(* Logix 5000 project; controller PLC_MCC1201_220AP1 vendor 1 type 14 code 164 rev 35.11; software revision 35.00; part 10 of 25 *)
(* tags used below, declared in another part *)
   TMP_rDummy : REAL;
   TMP_rTarget : REAL;
   TMP_xDummy : BOOL;
   B3 : DINT[102];
   GP_OB_InitializeMain : GP_OB_Initialize;
   HMI_Alarm_Reset : BOOL;   // HMI_Alarm_Reset
   HMI_MAN_CMD_WR : UDT_MAN_CMD_WR;
   LEHR_SPEED : ALIAS FOR N60[1];
   M225 : MAC_EMERGENCYXCUT;
   M225_HMW : MAC_EMERGENCYXCUT_HMW;
   M225_M1_DR : AXIS_CIP_DRIVE;
   M225_OUT_MOTION : MAC_EMERGENCYXCUT_OUT_MOTION;
   M2xx_CONVEYOR : MAC_CONVEYOR[20];
   M2xx_CONVEYOR_IN_MOTION : MAC_CONVEYOR_IN_MOTION[20];
   M2xx_CONVEYOR_OUT_MOTION : MAC_CONVEYOR_OUT_MOTION[20];
   M301_M1_DR : AXIS_CIP_DRIVE;
   M301_M2_DR : AXIS_CIP_DRIVE;
   TMP_dDirection : DINT;
   TMP_rAcc : REAL;
   TMP_rDec : REAL;
   TMP_rSpeed : REAL;
   TMP_xAlwaysOFF : BOOL;
   TMP_xRun : BOOL;
   Z200_UPS : ZONE_UPS;
(* CommandLogic, continued *)

ROUTINE M225_EmergencyCut_Outputs   (* ladder *)
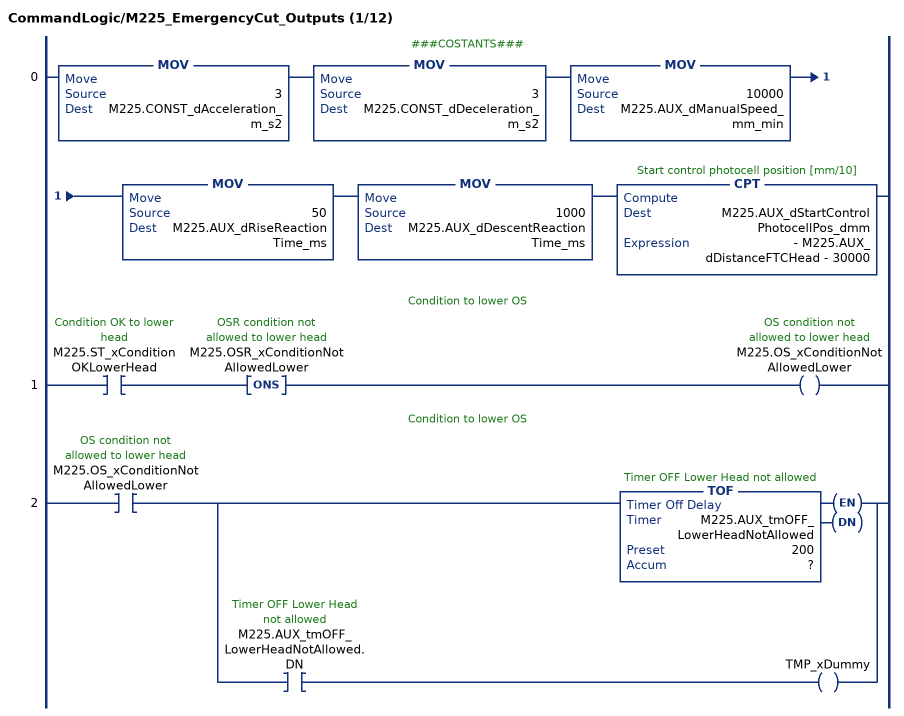
   // ###COSTANTS###
   0: MOV(3,M225.CONST_dAcceleration_m_s2)MOV(3,M225.CONST_dDeceleration_m_s2)MOV(10000,M225.AUX_dManualSpeed_mm_min)MOV(50,M225.AUX_dRiseReactionTime_ms)MOV(1000,M225.AUX_dDescentReactionTime_ms)CPT(M225.AUX_dStartControlPhotocellPos_dmm,- M225.AUX_dDistanceFTCHead - 30000);
   // Condition to lower OS
   1: XIC(M225.ST_xConditionOKLowerHead)ONS(M225.OSR_xConditionNotAllowedLower)OTE(M225.OS_xConditionNotAllowedLower);
   // Condition to lower OS
   2: XIC(M225.OS_xConditionNotAllowedLower)[TOF(M225.AUX_tmOFF_LowerHeadNotAllowed,?,?) ,XIC(M225.AUX_tmOFF_LowerHeadNotAllowed.DN) OTE(TMP_xDummy) ];
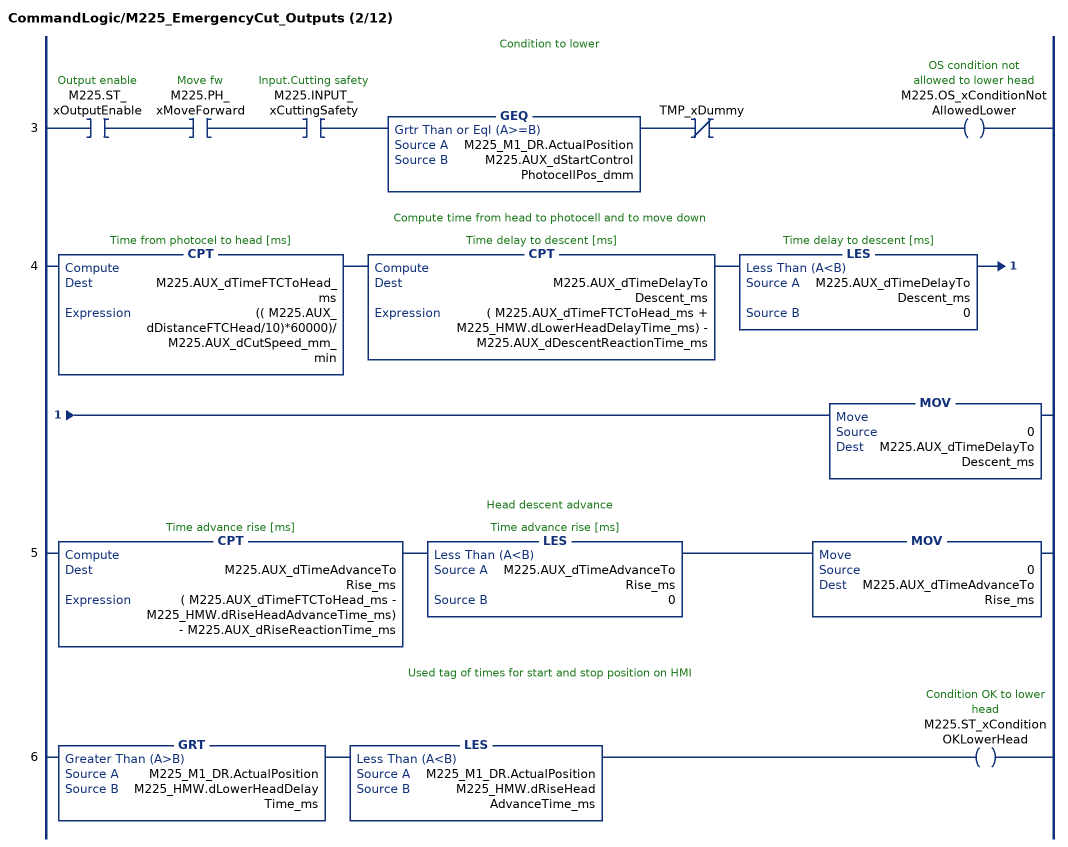
   // Condition to lower
   3: XIC(M225.ST_xOutputEnable)XIC(M225.PH_xMoveForward)XIC(M225.INPUT_xCuttingSafety)GEQ(M225_M1_DR.ActualPosition,M225.AUX_dStartControlPhotocellPos_dmm)XIO(TMP_xDummy)OTE(M225.OS_xConditionNotAllowedLower);
   // Compute time from head to photocell and to move down
   4: CPT(M225.AUX_dTimeFTCToHead_ms,(( M225.AUX_dDistanceFTCHead/10)*60000)/ M225.AUX_dCutSpeed_mm_min)CPT(M225.AUX_dTimeDelayToDescent_ms,( M225.AUX_dTimeFTCToHead_ms + M225_HMW.dLowerHeadDelayTime_ms) - M225.AUX_dDescentReactionTime_ms)LES(M225.AUX_dTimeDelayToDescent_ms,0)MOV(0,M225.AUX_dTimeDelayToDescent_ms);
   // Head descent advance
   5: CPT(M225.AUX_dTimeAdvanceToRise_ms,( M225.AUX_dTimeFTCToHead_ms - M225_HMW.dRiseHeadAdvanceTime_ms) - M225.AUX_dRiseReactionTime_ms)LES(M225.AUX_dTimeAdvanceToRise_ms,0)MOV(0,M225.AUX_dTimeAdvanceToRise_ms);
   // Used tag of times for start and stop position on HMI
   6: GRT(M225_M1_DR.ActualPosition,M225_HMW.dLowerHeadDelayTime_ms)LES(M225_M1_DR.ActualPosition,M225_HMW.dRiseHeadAdvanceTime_ms)OTE(M225.ST_xConditionOKLowerHead);
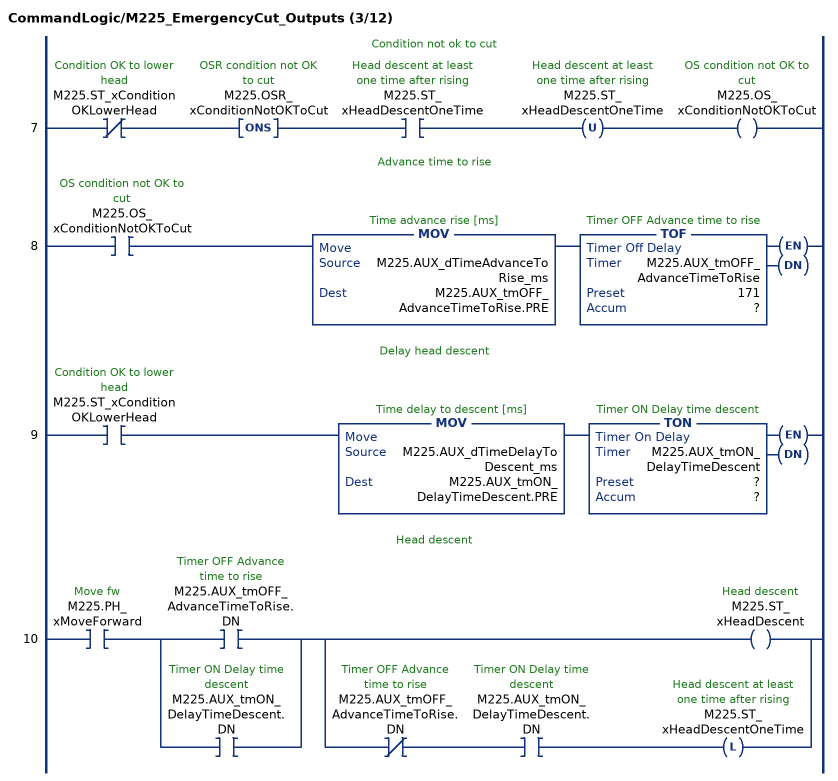
   // Condition not ok to cut
   7: XIO(M225.ST_xConditionOKLowerHead)ONS(M225.OSR_xConditionNotOKToCut)XIC(M225.ST_xHeadDescentOneTime)OTU(M225.ST_xHeadDescentOneTime)OTE(M225.OS_xConditionNotOKToCut);
   // Advance time to rise
   8: XIC(M225.OS_xConditionNotOKToCut)MOV(M225.AUX_dTimeAdvanceToRise_ms,M225.AUX_tmOFF_AdvanceTimeToRise.PRE)TOF(M225.AUX_tmOFF_AdvanceTimeToRise,?,?);
   // Delay head descent
   9: XIC(M225.ST_xConditionOKLowerHead)MOV(M225.AUX_dTimeDelayToDescent_ms,M225.AUX_tmON_DelayTimeDescent.PRE)TON(M225.AUX_tmON_DelayTimeDescent,?,?);
   // Head descent
   10: XIC(M225.PH_xMoveForward)[XIC(M225.AUX_tmOFF_AdvanceTimeToRise.DN) ,XIC(M225.AUX_tmON_DelayTimeDescent.DN) ][OTE(M225.ST_xHeadDescent) ,XIO(M225.AUX_tmOFF_AdvanceTimeToRise.DN) XIC(M225.AUX_tmON_DelayTimeDescent.DN) OTL(M225.ST_xHeadDescentOneTime) ];
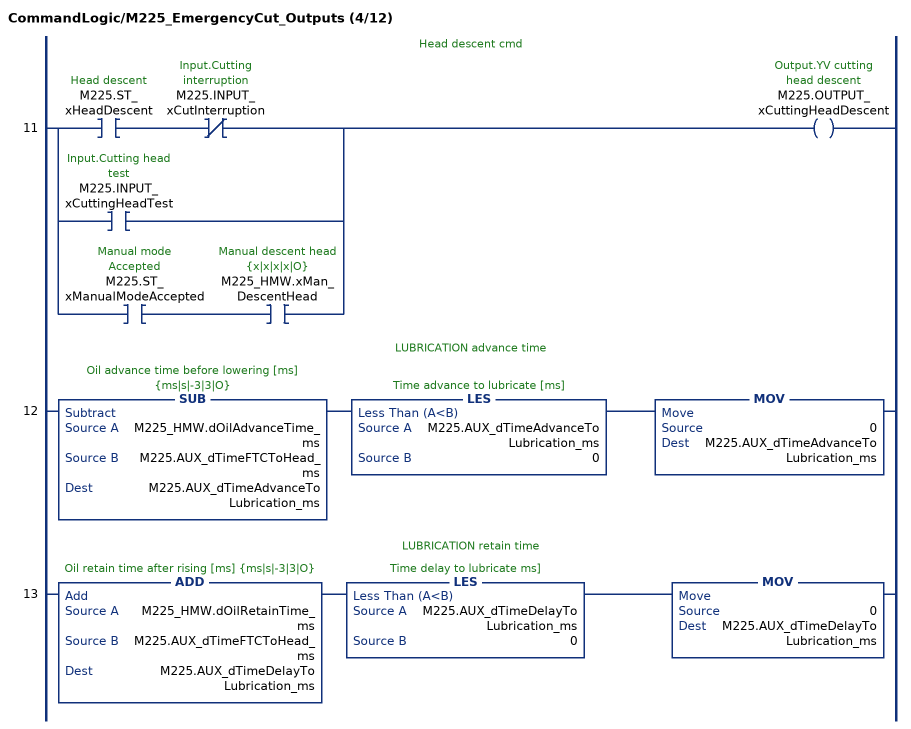
   // Head descent cmd
   11: [XIC(M225.ST_xHeadDescent) XIO(M225.INPUT_xCutInterruption) ,XIC(M225.INPUT_xCuttingHeadTest) ,XIC(M225.ST_xManualModeAccepted) XIC(M225_HMW.xMan_DescentHead) ]OTE(M225.OUTPUT_xCuttingHeadDescent);
   // LUBRICATION advance time
   12: SUB(M225_HMW.dOilAdvanceTime_ms,M225.AUX_dTimeFTCToHead_ms,M225.AUX_dTimeAdvanceToLubrication_ms)LES(M225.AUX_dTimeAdvanceToLubrication_ms,0)MOV(0,M225.AUX_dTimeAdvanceToLubrication_ms);
   // LUBRICATION retain time
   13: ADD(M225_HMW.dOilRetainTime_ms,M225.AUX_dTimeFTCToHead_ms,M225.AUX_dTimeDelayToLubrication_ms)LES(M225.AUX_dTimeDelayToLubrication_ms,0)MOV(0,M225.AUX_dTimeDelayToLubrication_ms);
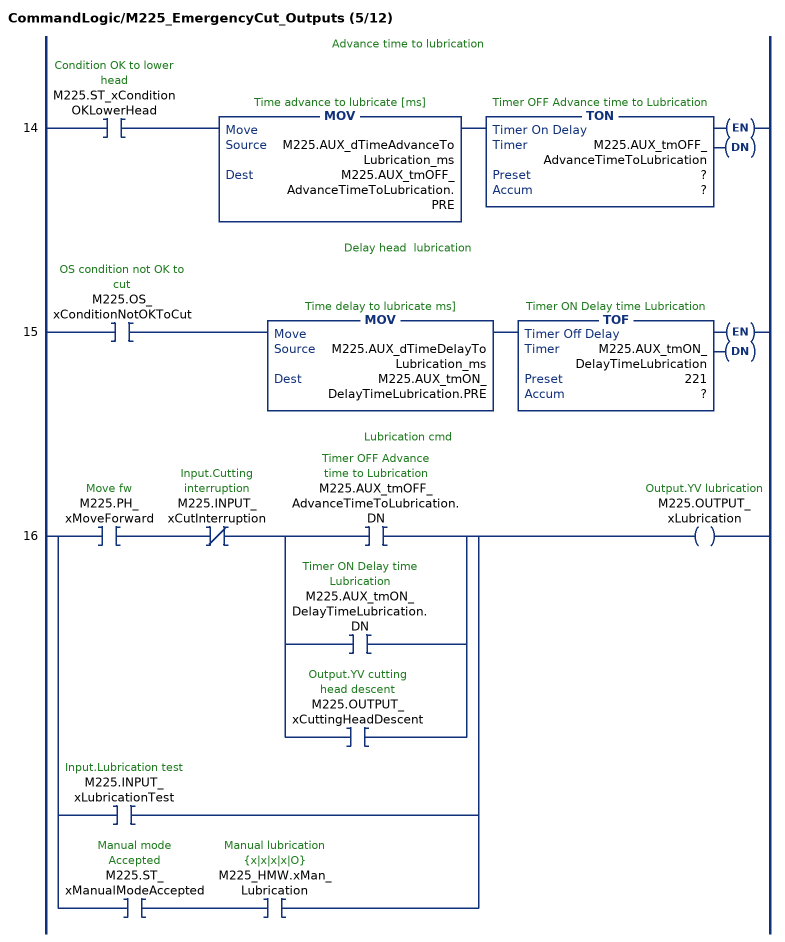
   // Advance time to lubrication
   14: XIC(M225.ST_xConditionOKLowerHead)MOV(M225.AUX_dTimeAdvanceToLubrication_ms,M225.AUX_tmOFF_AdvanceTimeToLubrication.PRE)TON(M225.AUX_tmOFF_AdvanceTimeToLubrication,?,?);
   // Delay head  lubrication
   15: XIC(M225.OS_xConditionNotOKToCut)MOV(M225.AUX_dTimeDelayToLubrication_ms,M225.AUX_tmON_DelayTimeLubrication.PRE)TOF(M225.AUX_tmON_DelayTimeLubrication,?,?);
   // Lubrication cmd
   16: [XIC(M225.PH_xMoveForward) XIO(M225.INPUT_xCutInterruption) [XIC(M225.AUX_tmOFF_AdvanceTimeToLubrication.DN) ,XIC(M225.AUX_tmON_DelayTimeLubrication.DN) ,XIC(M225.OUTPUT_xCuttingHeadDescent) ] ,XIC(M225.INPUT_xLubricationTest) ,XIC(M225.ST_xManualModeAccepted) XIC(M225_HMW.xMan_Lubrication) ]OTE(M225.OUTPUT_xLubrication);
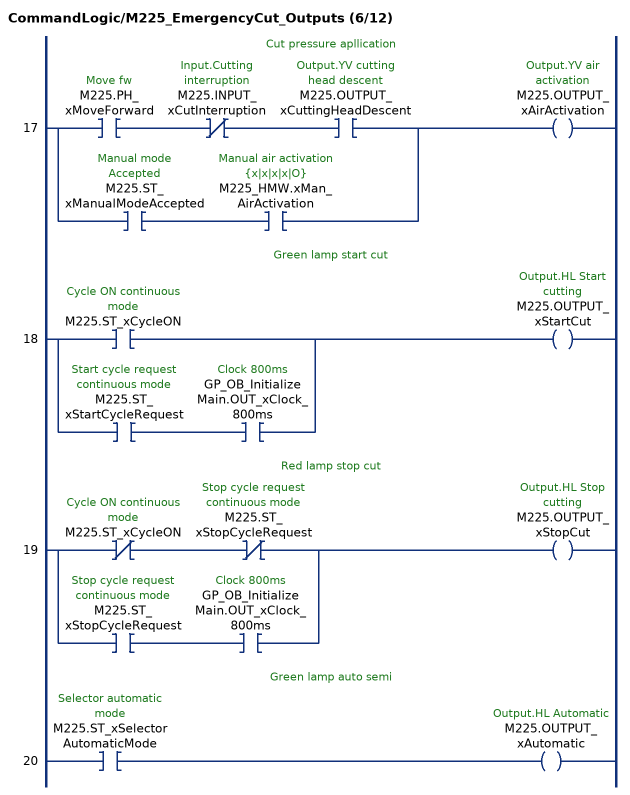
   // Cut pressure apllication
   17: [XIC(M225.PH_xMoveForward) XIO(M225.INPUT_xCutInterruption) XIC(M225.OUTPUT_xCuttingHeadDescent) ,XIC(M225.ST_xManualModeAccepted) XIC(M225_HMW.xMan_AirActivation) ]OTE(M225.OUTPUT_xAirActivation);
   // Green lamp start cut
   18: [XIC(M225.ST_xCycleON) ,XIC(M225.ST_xStartCycleRequest) XIC(GP_OB_InitializeMain.OUT_xClock_800ms) ]OTE(M225.OUTPUT_xStartCut);
   // Red lamp stop cut
   19: [XIO(M225.ST_xCycleON) XIO(M225.ST_xStopCycleRequest) ,XIC(M225.ST_xStopCycleRequest) XIC(GP_OB_InitializeMain.OUT_xClock_800ms) ]OTE(M225.OUTPUT_xStopCut);
   // Green lamp auto semi
   20: XIC(M225.ST_xSelectorAutomaticMode)OTE(M225.OUTPUT_xAutomatic);
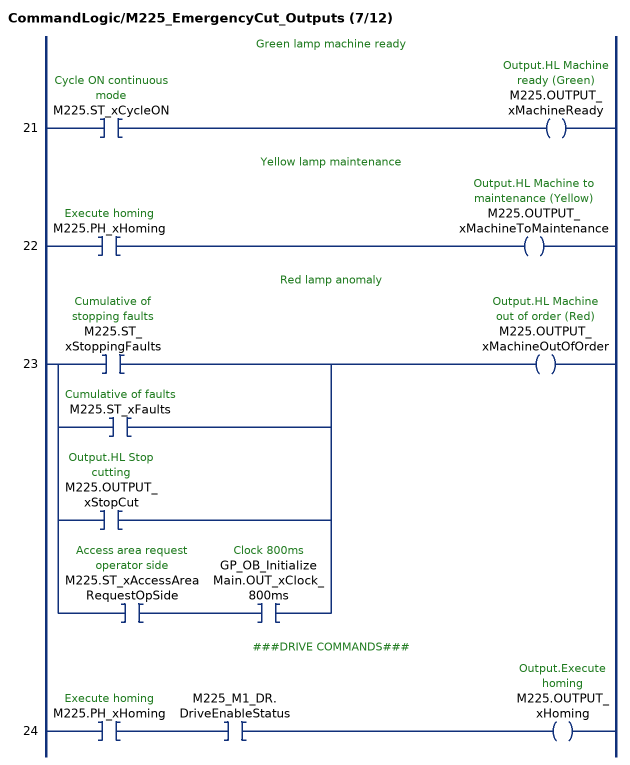
   // Green lamp machine ready
   21: XIC(M225.ST_xCycleON)OTE(M225.OUTPUT_xMachineReady);
   // Yellow lamp maintenance
   22: XIC(M225.PH_xHoming)OTE(M225.OUTPUT_xMachineToMaintenance);
   // Red lamp anomaly
   23: [XIC(M225.ST_xStoppingFaults) ,XIC(M225.ST_xFaults) ,XIC(M225.OUTPUT_xStopCut) ,XIC(M225.ST_xAccessAreaRequestOpSide) XIC(GP_OB_InitializeMain.OUT_xClock_800ms) ]OTE(M225.OUTPUT_xMachineOutOfOrder);
   // ###DRIVE COMMANDS###
   24: XIC(M225.PH_xHoming)XIC(M225_M1_DR.DriveEnableStatus)OTE(M225.OUTPUT_xHoming);
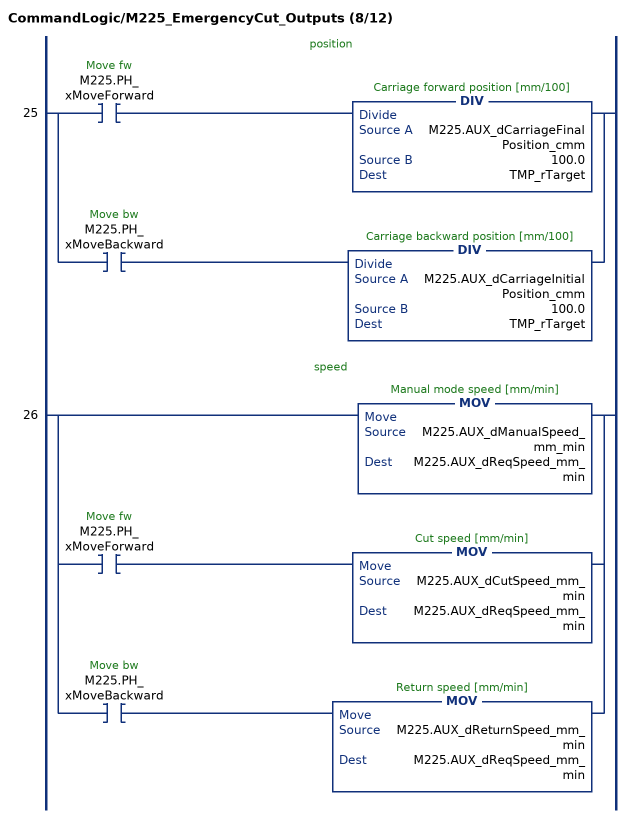
   // position
   25: [XIC(M225.PH_xMoveForward) DIV(M225.AUX_dCarriageFinalPosition_cmm,100.0,TMP_rTarget) ,XIC(M225.PH_xMoveBackward) DIV(M225.AUX_dCarriageInitialPosition_cmm,100.0,TMP_rTarget) ];
   // speed
   26: [MOV(M225.AUX_dManualSpeed_mm_min,M225.AUX_dReqSpeed_mm_min) ,XIC(M225.PH_xMoveForward) MOV(M225.AUX_dCutSpeed_mm_min,M225.AUX_dReqSpeed_mm_min) ,XIC(M225.PH_xMoveBackward) MOV(M225.AUX_dReturnSpeed_mm_min,M225.AUX_dReqSpeed_mm_min) ];
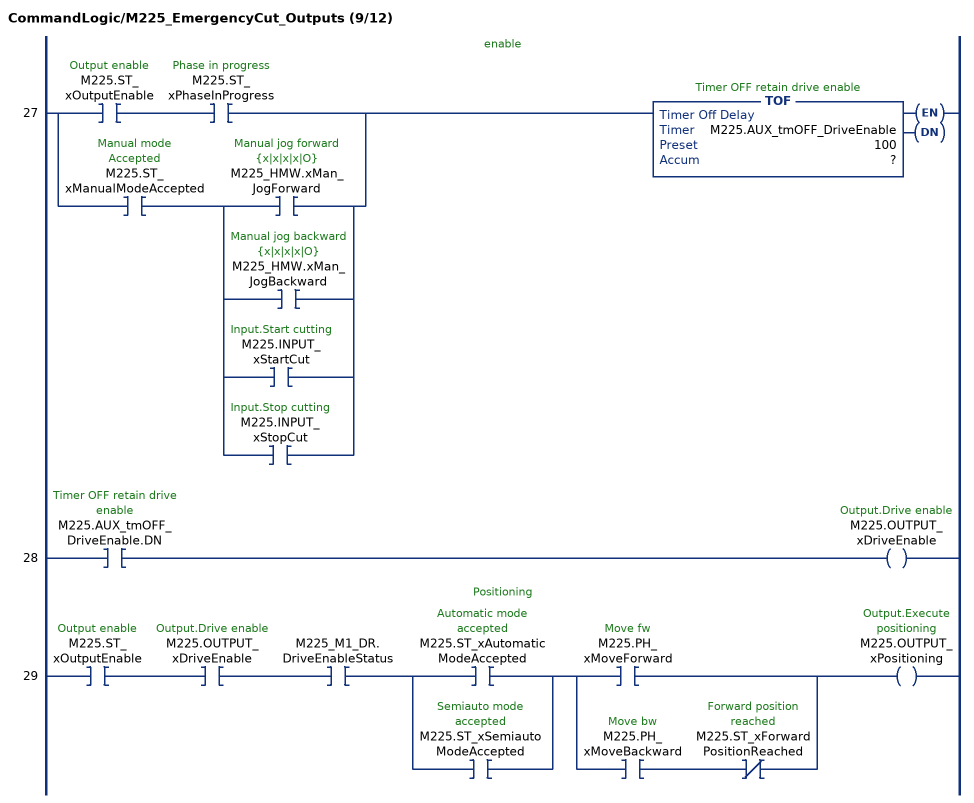
   // enable
   27: [XIC(M225.ST_xOutputEnable) XIC(M225.ST_xPhaseInProgress) ,XIC(M225.ST_xManualModeAccepted) [XIC(M225_HMW.xMan_JogForward) ,XIC(M225_HMW.xMan_JogBackward) ,XIC(M225.INPUT_xStartCut) ,XIC(M225.INPUT_xStopCut) ] ]TOF(M225.AUX_tmOFF_DriveEnable,?,?);
   28: XIC(M225.AUX_tmOFF_DriveEnable.DN)OTE(M225.OUTPUT_xDriveEnable);
   // Positioning
   29: XIC(M225.ST_xOutputEnable)XIC(M225.OUTPUT_xDriveEnable)XIC(M225_M1_DR.DriveEnableStatus)[XIC(M225.ST_xAutomaticModeAccepted) ,XIC(M225.ST_xSemiautoModeAccepted) ][XIC(M225.PH_xMoveForward) ,XIC(M225.PH_xMoveBackward) XIO(M225.ST_xForwardPositionReached) ]OTE(M225.OUTPUT_xPositioning);
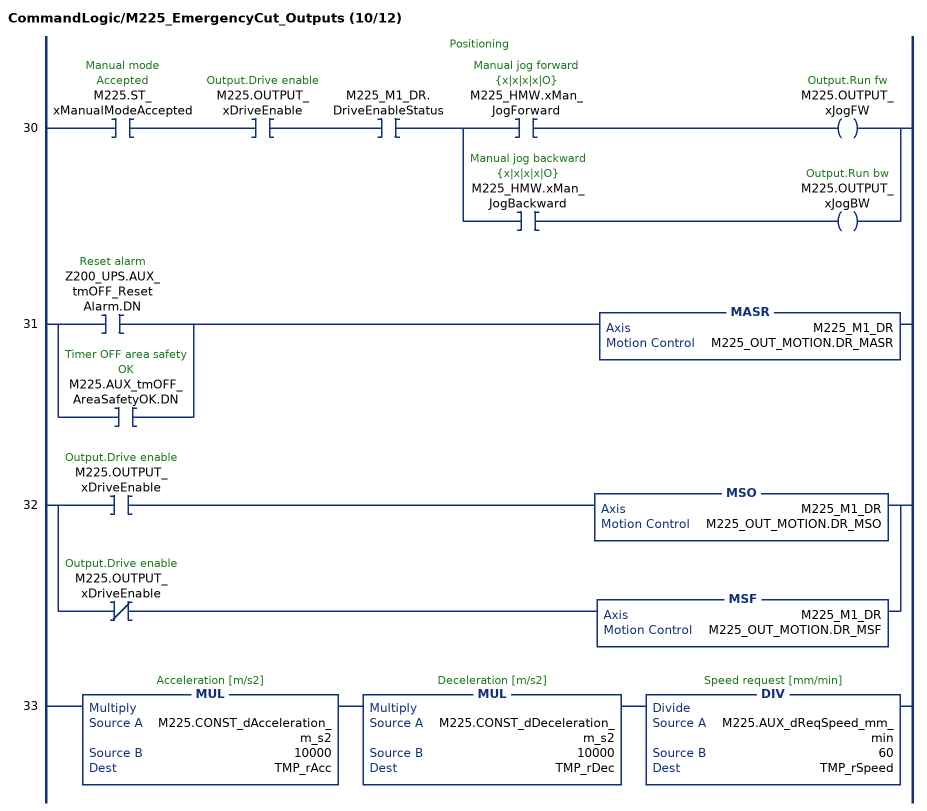
   // Positioning
   30: XIC(M225.ST_xManualModeAccepted)XIC(M225.OUTPUT_xDriveEnable)XIC(M225_M1_DR.DriveEnableStatus)[XIC(M225_HMW.xMan_JogForward) OTE(M225.OUTPUT_xJogFW) ,XIC(M225_HMW.xMan_JogBackward) OTE(M225.OUTPUT_xJogBW) ];
   31: [XIC(Z200_UPS.AUX_tmOFF_ResetAlarm.DN) ,XIC(M225.AUX_tmOFF_AreaSafetyOK.DN) ]MASR(M225_M1_DR,M225_OUT_MOTION.DR_MASR);
   32: [XIC(M225.OUTPUT_xDriveEnable) MSO(M225_M1_DR,M225_OUT_MOTION.DR_MSO) ,XIO(M225.OUTPUT_xDriveEnable) MSF(M225_M1_DR,M225_OUT_MOTION.DR_MSF) ];
   33: MUL(M225.CONST_dAcceleration_m_s2,10000,TMP_rAcc)MUL(M225.CONST_dDeceleration_m_s2,10000,TMP_rDec)DIV(M225.AUX_dReqSpeed_mm_min,60,TMP_rSpeed);
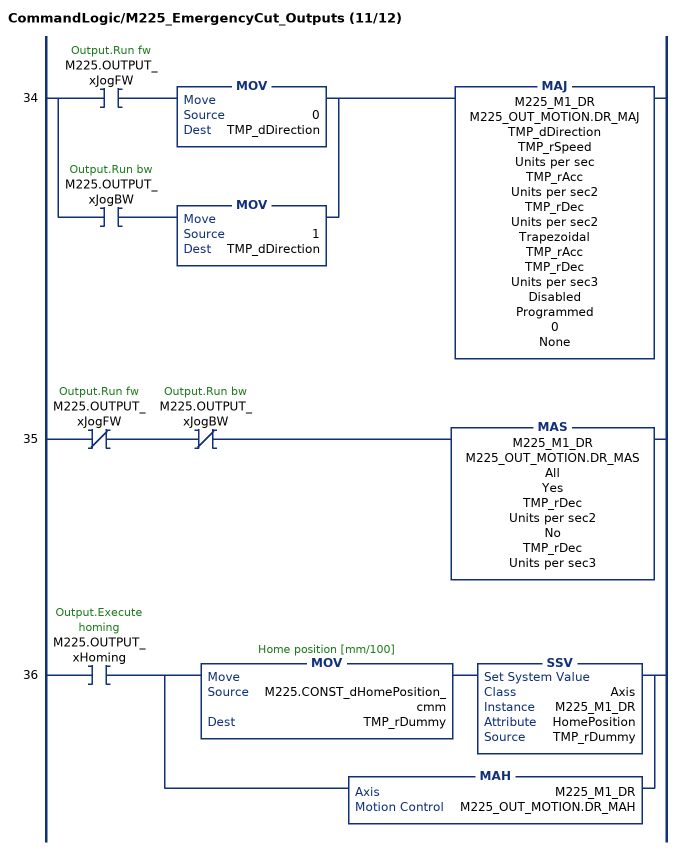
   34: [XIC(M225.OUTPUT_xJogFW) MOV(0,TMP_dDirection) ,XIC(M225.OUTPUT_xJogBW) MOV(1,TMP_dDirection) ]MAJ(M225_M1_DR,M225_OUT_MOTION.DR_MAJ,TMP_dDirection,TMP_rSpeed,Units per sec,TMP_rAcc,Units per sec2,TMP_rDec,Units per sec2,Trapezoidal,TMP_rAcc,TMP_rDec,Units per sec3,Disabled,Programmed,0,None);
   35: XIO(M225.OUTPUT_xJogFW)XIO(M225.OUTPUT_xJogBW)MAS(M225_M1_DR,M225_OUT_MOTION.DR_MAS,All,Yes,TMP_rDec,Units per sec2,No,TMP_rDec,Units per sec3);
   36: XIC(M225.OUTPUT_xHoming)[MOV(M225.CONST_dHomePosition_cmm,TMP_rDummy) SSV(Axis,M225_M1_DR,HomePosition,TMP_rDummy) ,MAH(M225_M1_DR,M225_OUT_MOTION.DR_MAH) ];
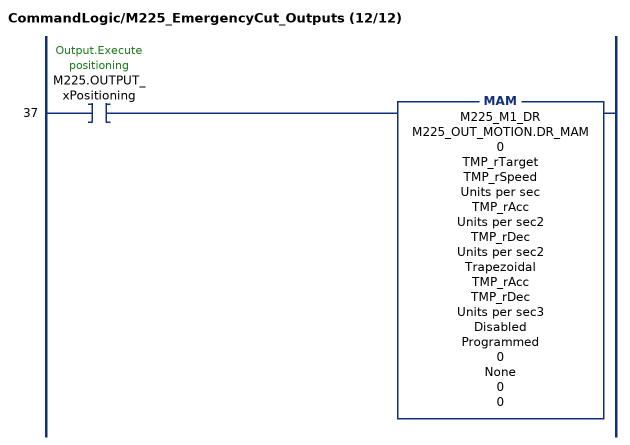
   37: XIC(M225.OUTPUT_xPositioning)MAM(M225_M1_DR,M225_OUT_MOTION.DR_MAM,0,TMP_rTarget,TMP_rSpeed,Units per sec,TMP_rAcc,Units per sec2,TMP_rDec,Units per sec2,Trapezoidal,TMP_rAcc,TMP_rDec,Units per sec3,Disabled,Programmed,0,None,0,0);
END_ROUTINE

ROUTINE M301M1_Conveyor_Motion_Output   (* ladder *)
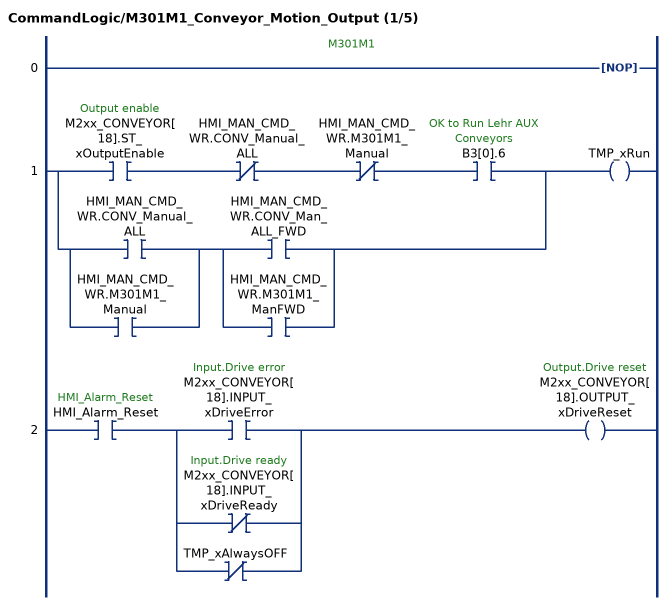
   // M301M1
   0: NOP();
   1: [XIC(M2xx_CONVEYOR[18].ST_xOutputEnable) XIO(HMI_MAN_CMD_WR.CONV_Manual_ALL) XIO(HMI_MAN_CMD_WR.M301M1_Manual) XIC(B3[0].6) ,[XIC(HMI_MAN_CMD_WR.CONV_Manual_ALL) ,XIC(HMI_MAN_CMD_WR.M301M1_Manual) ] [XIC(HMI_MAN_CMD_WR.CONV_Man_ALL_FWD) ,XIC(HMI_MAN_CMD_WR.M301M1_ManFWD) ] ]OTE(TMP_xRun);
   2: XIC(HMI_Alarm_Reset)[XIC(M2xx_CONVEYOR[18].INPUT_xDriveError) ,XIO(M2xx_CONVEYOR[18].INPUT_xDriveReady) ,XIO(TMP_xAlwaysOFF) ]OTE(M2xx_CONVEYOR[18].OUTPUT_xDriveReset);
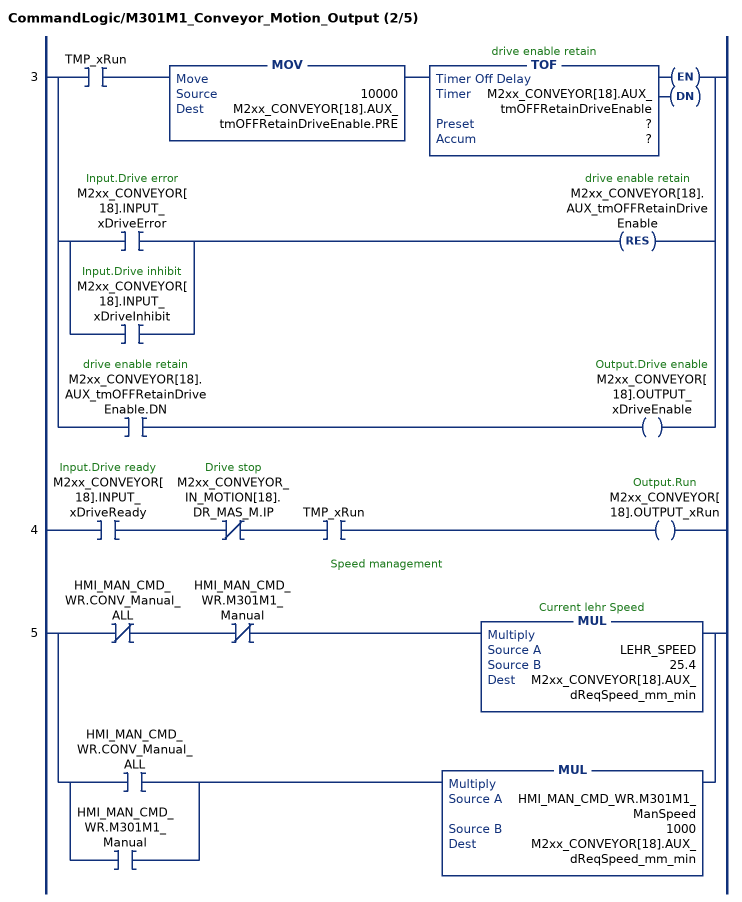
   3: [XIC(TMP_xRun) MOV(10000,M2xx_CONVEYOR[18].AUX_tmOFFRetainDriveEnable.PRE) TOF(M2xx_CONVEYOR[18].AUX_tmOFFRetainDriveEnable,?,?) ,[XIC(M2xx_CONVEYOR[18].INPUT_xDriveError) ,XIC(M2xx_CONVEYOR[18].INPUT_xDriveInhibit) ] RES(M2xx_CONVEYOR[18].AUX_tmOFFRetainDriveEnable) ,XIC(M2xx_CONVEYOR[18].AUX_tmOFFRetainDriveEnable.DN) OTE(M2xx_CONVEYOR[18].OUTPUT_xDriveEnable) ];
   4: XIC(M2xx_CONVEYOR[18].INPUT_xDriveReady)XIO(M2xx_CONVEYOR_IN_MOTION[18].DR_MAS_M.IP)XIC(TMP_xRun)OTE(M2xx_CONVEYOR[18].OUTPUT_xRun);
   // Speed management
   5: [XIO(HMI_MAN_CMD_WR.CONV_Manual_ALL) XIO(HMI_MAN_CMD_WR.M301M1_Manual) MUL(LEHR_SPEED,25.4,M2xx_CONVEYOR[18].AUX_dReqSpeed_mm_min) ,[XIC(HMI_MAN_CMD_WR.CONV_Manual_ALL) ,XIC(HMI_MAN_CMD_WR.M301M1_Manual) ] MUL(HMI_MAN_CMD_WR.M301M1_ManSpeed,1000,M2xx_CONVEYOR[18].AUX_dReqSpeed_mm_min) ];
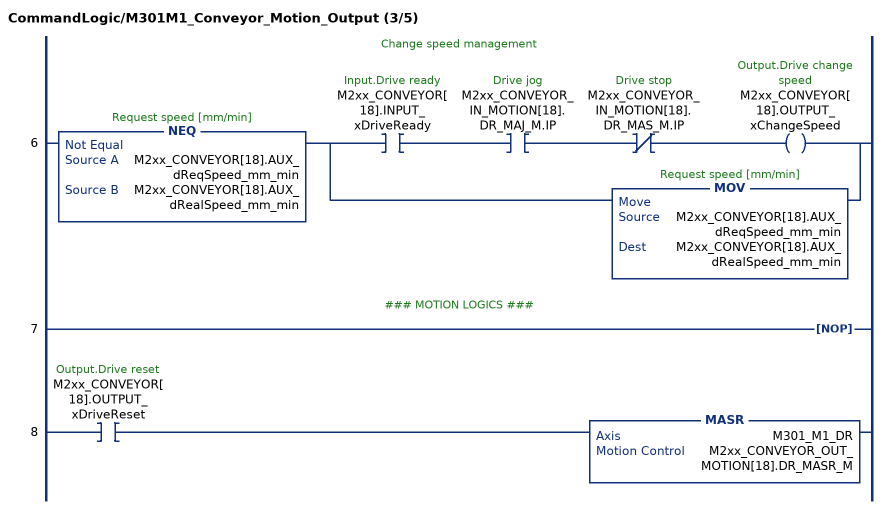
   // Change speed management
   6: NEQ(M2xx_CONVEYOR[18].AUX_dReqSpeed_mm_min,M2xx_CONVEYOR[18].AUX_dRealSpeed_mm_min)[XIC(M2xx_CONVEYOR[18].INPUT_xDriveReady) XIC(M2xx_CONVEYOR_IN_MOTION[18].DR_MAJ_M.IP) XIO(M2xx_CONVEYOR_IN_MOTION[18].DR_MAS_M.IP) OTE(M2xx_CONVEYOR[18].OUTPUT_xChangeSpeed) ,MOV(M2xx_CONVEYOR[18].AUX_dReqSpeed_mm_min,M2xx_CONVEYOR[18].AUX_dRealSpeed_mm_min) ];
   // ### MOTION LOGICS ###
   7: NOP();
   8: XIC(M2xx_CONVEYOR[18].OUTPUT_xDriveReset)MASR(M301_M1_DR,M2xx_CONVEYOR_OUT_MOTION[18].DR_MASR_M);
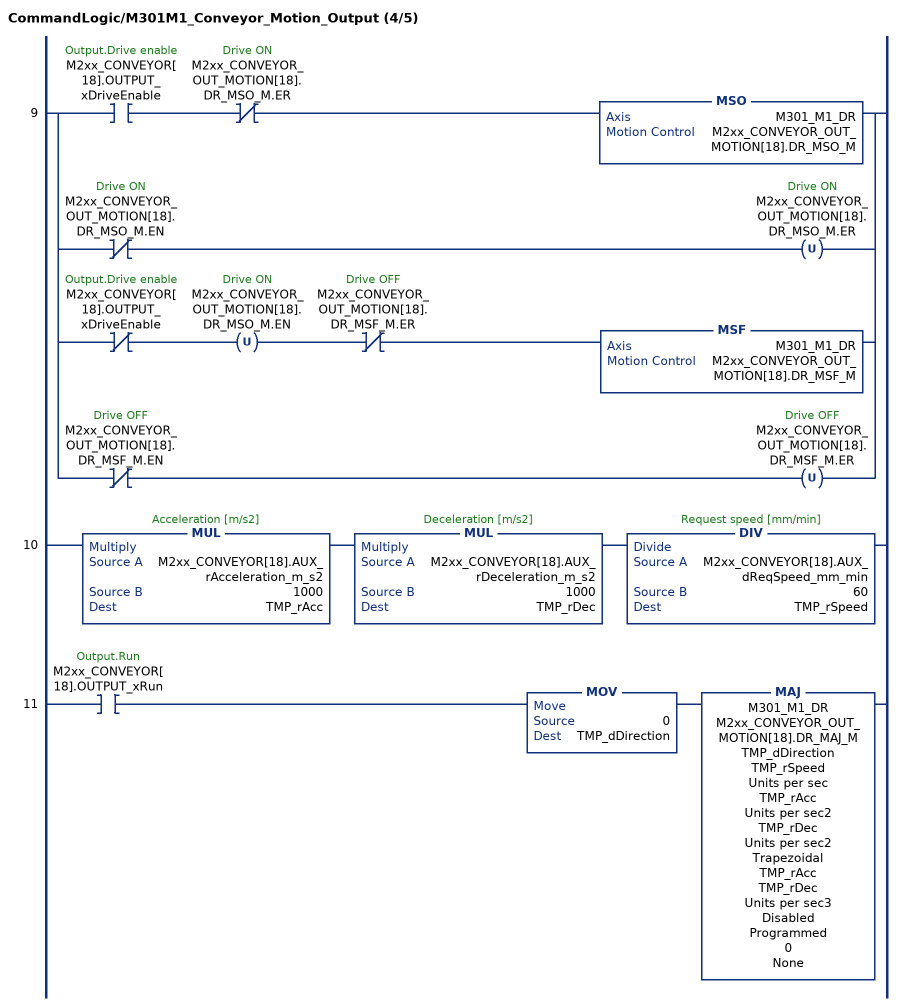
   9: [XIC(M2xx_CONVEYOR[18].OUTPUT_xDriveEnable) XIO(M2xx_CONVEYOR_OUT_MOTION[18].DR_MSO_M.ER) MSO(M301_M1_DR,M2xx_CONVEYOR_OUT_MOTION[18].DR_MSO_M) ,XIO(M2xx_CONVEYOR_OUT_MOTION[18].DR_MSO_M.EN) OTU(M2xx_CONVEYOR_OUT_MOTION[18].DR_MSO_M.ER) ,XIO(M2xx_CONVEYOR[18].OUTPUT_xDriveEnable) OTU(M2xx_CONVEYOR_OUT_MOTION[18].DR_MSO_M.EN) XIO(M2xx_CONVEYOR_OUT_MOTION[18].DR_MSF_M.ER) MSF(M301_M1_DR,M2xx_CONVEYOR_OUT_MOTION[18].DR_MSF_M) ,XIO(M2xx_CONVEYOR_OUT_MOTION[18].DR_MSF_M.EN) OTU(M2xx_CONVEYOR_OUT_MOTION[18].DR_MSF_M.ER) ];
   10: MUL(M2xx_CONVEYOR[18].AUX_rAcceleration_m_s2,1000,TMP_rAcc)MUL(M2xx_CONVEYOR[18].AUX_rDeceleration_m_s2,1000,TMP_rDec)DIV(M2xx_CONVEYOR[18].AUX_dReqSpeed_mm_min,60,TMP_rSpeed);
   11: XIC(M2xx_CONVEYOR[18].OUTPUT_xRun)MOV(0,TMP_dDirection)MAJ(M301_M1_DR,M2xx_CONVEYOR_OUT_MOTION[18].DR_MAJ_M,TMP_dDirection,TMP_rSpeed,Units per sec,TMP_rAcc,Units per sec2,TMP_rDec,Units per sec2,Trapezoidal,TMP_rAcc,TMP_rDec,Units per sec3,Disabled,Programmed,0,None);
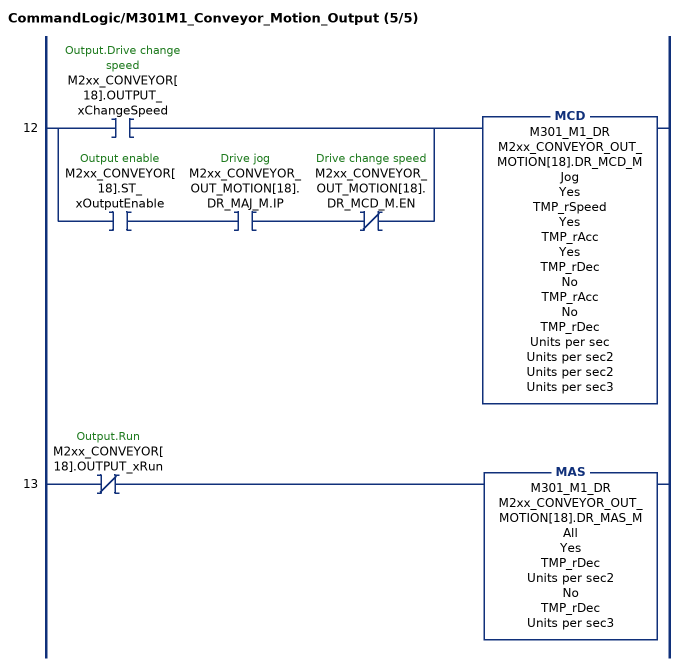
   12: [XIC(M2xx_CONVEYOR[18].OUTPUT_xChangeSpeed) ,XIC(M2xx_CONVEYOR[18].ST_xOutputEnable) XIC(M2xx_CONVEYOR_OUT_MOTION[18].DR_MAJ_M.IP) XIO(M2xx_CONVEYOR_OUT_MOTION[18].DR_MCD_M.EN) ]MCD(M301_M1_DR,M2xx_CONVEYOR_OUT_MOTION[18].DR_MCD_M,Jog,Yes,TMP_rSpeed,Yes,TMP_rAcc,Yes,TMP_rDec,No,TMP_rAcc,No,TMP_rDec,Units per sec,Units per sec2,Units per sec2,Units per sec3);
   13: XIO(M2xx_CONVEYOR[18].OUTPUT_xRun)MAS(M301_M1_DR,M2xx_CONVEYOR_OUT_MOTION[18].DR_MAS_M,All,Yes,TMP_rDec,Units per sec2,No,TMP_rDec,Units per sec3);
END_ROUTINE

ROUTINE M301M2_Conveyor_Motion_Output   (* ladder *)
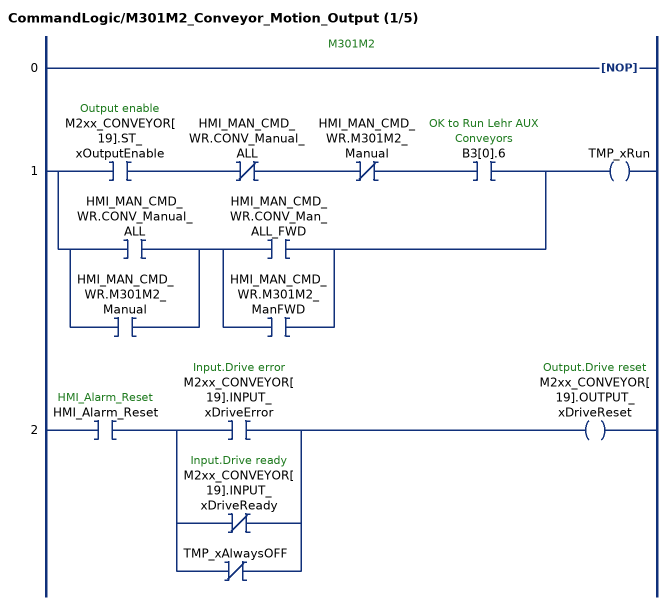
   // M301M2
   0: NOP();
   1: [XIC(M2xx_CONVEYOR[19].ST_xOutputEnable) XIO(HMI_MAN_CMD_WR.CONV_Manual_ALL) XIO(HMI_MAN_CMD_WR.M301M2_Manual) XIC(B3[0].6) ,[XIC(HMI_MAN_CMD_WR.CONV_Manual_ALL) ,XIC(HMI_MAN_CMD_WR.M301M2_Manual) ] [XIC(HMI_MAN_CMD_WR.CONV_Man_ALL_FWD) ,XIC(HMI_MAN_CMD_WR.M301M2_ManFWD) ] ]OTE(TMP_xRun);
   2: XIC(HMI_Alarm_Reset)[XIC(M2xx_CONVEYOR[19].INPUT_xDriveError) ,XIO(M2xx_CONVEYOR[19].INPUT_xDriveReady) ,XIO(TMP_xAlwaysOFF) ]OTE(M2xx_CONVEYOR[19].OUTPUT_xDriveReset);
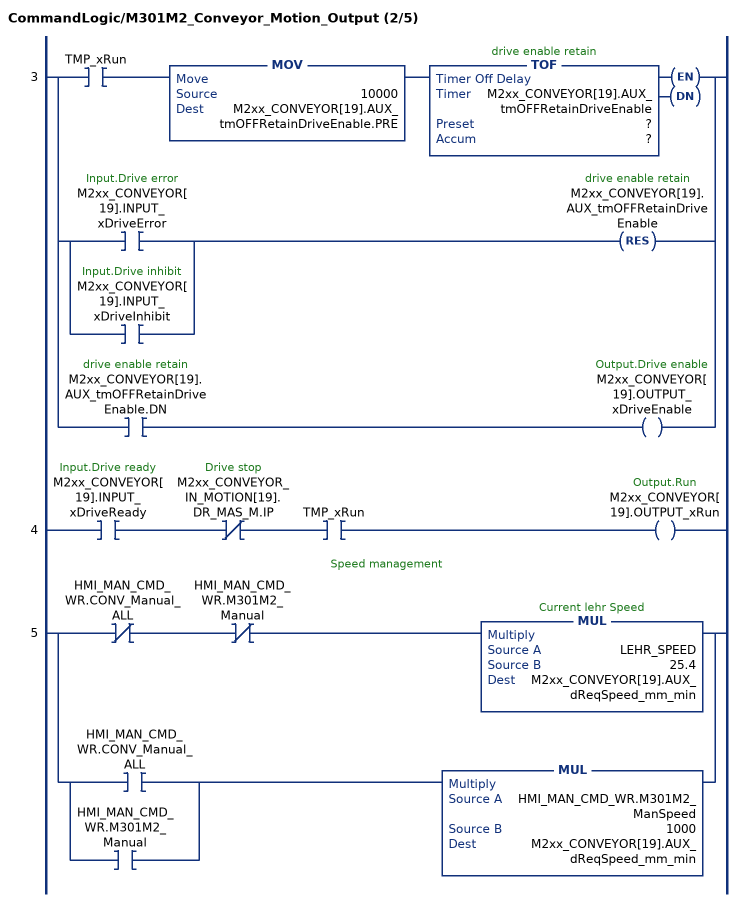
   3: [XIC(TMP_xRun) MOV(10000,M2xx_CONVEYOR[19].AUX_tmOFFRetainDriveEnable.PRE) TOF(M2xx_CONVEYOR[19].AUX_tmOFFRetainDriveEnable,?,?) ,[XIC(M2xx_CONVEYOR[19].INPUT_xDriveError) ,XIC(M2xx_CONVEYOR[19].INPUT_xDriveInhibit) ] RES(M2xx_CONVEYOR[19].AUX_tmOFFRetainDriveEnable) ,XIC(M2xx_CONVEYOR[19].AUX_tmOFFRetainDriveEnable.DN) OTE(M2xx_CONVEYOR[19].OUTPUT_xDriveEnable) ];
   4: XIC(M2xx_CONVEYOR[19].INPUT_xDriveReady)XIO(M2xx_CONVEYOR_IN_MOTION[19].DR_MAS_M.IP)XIC(TMP_xRun)OTE(M2xx_CONVEYOR[19].OUTPUT_xRun);
   // Speed management
   5: [XIO(HMI_MAN_CMD_WR.CONV_Manual_ALL) XIO(HMI_MAN_CMD_WR.M301M2_Manual) MUL(LEHR_SPEED,25.4,M2xx_CONVEYOR[19].AUX_dReqSpeed_mm_min) ,[XIC(HMI_MAN_CMD_WR.CONV_Manual_ALL) ,XIC(HMI_MAN_CMD_WR.M301M2_Manual) ] MUL(HMI_MAN_CMD_WR.M301M2_ManSpeed,1000,M2xx_CONVEYOR[19].AUX_dReqSpeed_mm_min) ];
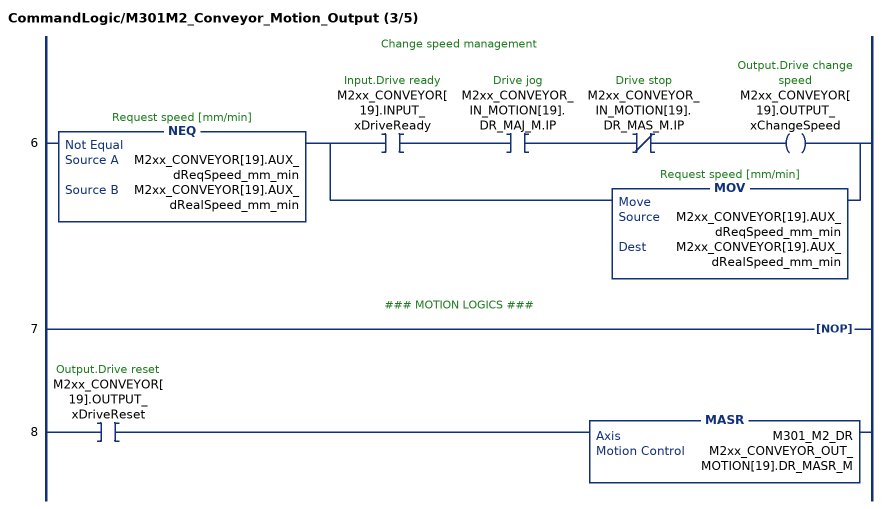
   // Change speed management
   6: NEQ(M2xx_CONVEYOR[19].AUX_dReqSpeed_mm_min,M2xx_CONVEYOR[19].AUX_dRealSpeed_mm_min)[XIC(M2xx_CONVEYOR[19].INPUT_xDriveReady) XIC(M2xx_CONVEYOR_IN_MOTION[19].DR_MAJ_M.IP) XIO(M2xx_CONVEYOR_IN_MOTION[19].DR_MAS_M.IP) OTE(M2xx_CONVEYOR[19].OUTPUT_xChangeSpeed) ,MOV(M2xx_CONVEYOR[19].AUX_dReqSpeed_mm_min,M2xx_CONVEYOR[19].AUX_dRealSpeed_mm_min) ];
   // ### MOTION LOGICS ###
   7: NOP();
   8: XIC(M2xx_CONVEYOR[19].OUTPUT_xDriveReset)MASR(M301_M2_DR,M2xx_CONVEYOR_OUT_MOTION[19].DR_MASR_M);
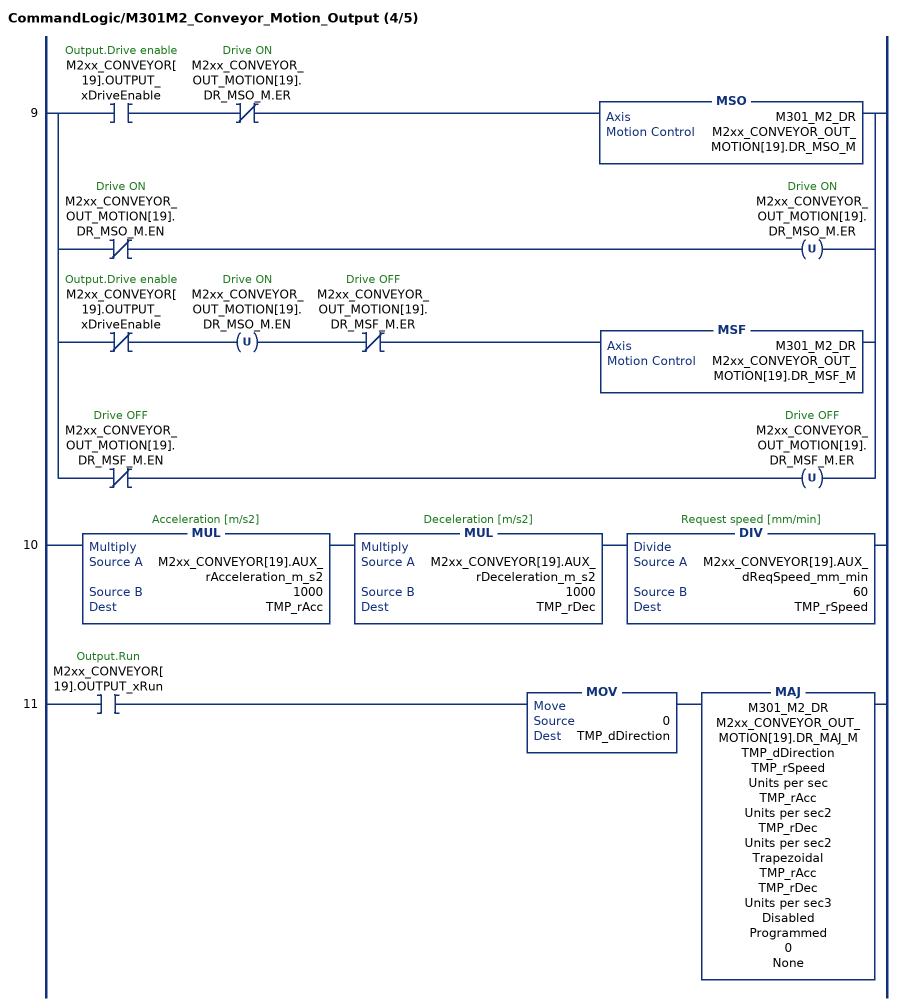
   9: [XIC(M2xx_CONVEYOR[19].OUTPUT_xDriveEnable) XIO(M2xx_CONVEYOR_OUT_MOTION[19].DR_MSO_M.ER) MSO(M301_M2_DR,M2xx_CONVEYOR_OUT_MOTION[19].DR_MSO_M) ,XIO(M2xx_CONVEYOR_OUT_MOTION[19].DR_MSO_M.EN) OTU(M2xx_CONVEYOR_OUT_MOTION[19].DR_MSO_M.ER) ,XIO(M2xx_CONVEYOR[19].OUTPUT_xDriveEnable) OTU(M2xx_CONVEYOR_OUT_MOTION[19].DR_MSO_M.EN) XIO(M2xx_CONVEYOR_OUT_MOTION[19].DR_MSF_M.ER) MSF(M301_M2_DR,M2xx_CONVEYOR_OUT_MOTION[19].DR_MSF_M) ,XIO(M2xx_CONVEYOR_OUT_MOTION[19].DR_MSF_M.EN) OTU(M2xx_CONVEYOR_OUT_MOTION[19].DR_MSF_M.ER) ];
   10: MUL(M2xx_CONVEYOR[19].AUX_rAcceleration_m_s2,1000,TMP_rAcc)MUL(M2xx_CONVEYOR[19].AUX_rDeceleration_m_s2,1000,TMP_rDec)DIV(M2xx_CONVEYOR[19].AUX_dReqSpeed_mm_min,60,TMP_rSpeed);
   11: XIC(M2xx_CONVEYOR[19].OUTPUT_xRun)MOV(0,TMP_dDirection)MAJ(M301_M2_DR,M2xx_CONVEYOR_OUT_MOTION[19].DR_MAJ_M,TMP_dDirection,TMP_rSpeed,Units per sec,TMP_rAcc,Units per sec2,TMP_rDec,Units per sec2,Trapezoidal,TMP_rAcc,TMP_rDec,Units per sec3,Disabled,Programmed,0,None);
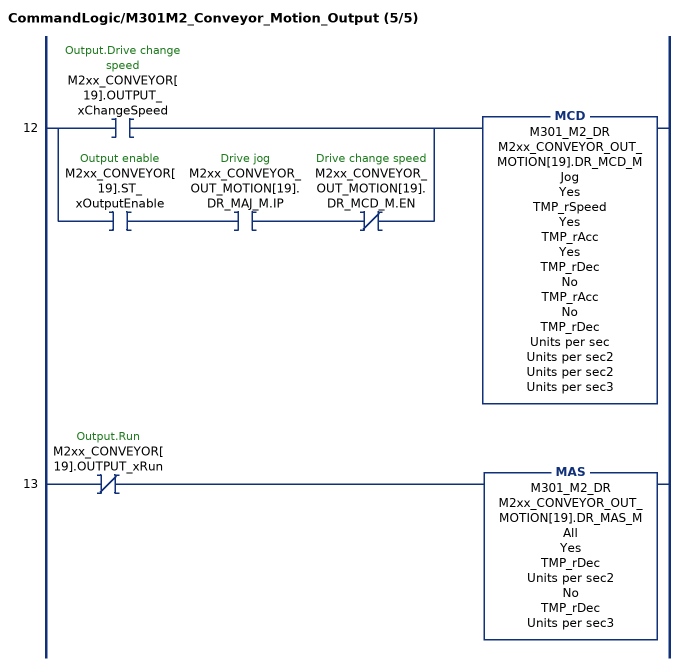
   12: [XIC(M2xx_CONVEYOR[19].OUTPUT_xChangeSpeed) ,XIC(M2xx_CONVEYOR[19].ST_xOutputEnable) XIC(M2xx_CONVEYOR_OUT_MOTION[19].DR_MAJ_M.IP) XIO(M2xx_CONVEYOR_OUT_MOTION[19].DR_MCD_M.EN) ]MCD(M301_M2_DR,M2xx_CONVEYOR_OUT_MOTION[19].DR_MCD_M,Jog,Yes,TMP_rSpeed,Yes,TMP_rAcc,Yes,TMP_rDec,No,TMP_rAcc,No,TMP_rDec,Units per sec,Units per sec2,Units per sec2,Units per sec3);
   13: XIO(M2xx_CONVEYOR[19].OUTPUT_xRun)MAS(M301_M2_DR,M2xx_CONVEYOR_OUT_MOTION[19].DR_MAS_M,All,Yes,TMP_rDec,Units per sec2,No,TMP_rDec,Units per sec3);
END_ROUTINE
